REGION Network 83
   RUNG wire#powerrail
      Move(in := "Carrier_44_G120DControlWord", out1 => "DB402_SDC_CARRIER_DRIVE_DATA".Drive_Data.CARRIER[44].Drive_Control)
      Move(in := "Carrier_44_G120DStatusWord", out1 => "DB402_SDC_CARRIER_DRIVE_DATA".Drive_Data.CARRIER[44].Drive_Status)
   END_RUNG
   // the same network as SCL:
   "DB402_SDC_CARRIER_DRIVE_DATA".Drive_Data.CARRIER[44].Drive_Control := "Carrier_44_G120DControlWord";
   "DB402_SDC_CARRIER_DRIVE_DATA".Drive_Data.CARRIER[44].Drive_Status := "Carrier_44_G120DStatusWord";
END_REGION

REGION Network 84
   RUNG wire#powerrail
      Move(in := "Carrier_44_SDCFaultCode", out1 => "DB_SDC_EMS_TA".EMS[44].TA[1].FAULT)
      wire#w1
      Move(in := "Carrier_44_SDCFaultCode", out1 => "EMS".Carrier[44].SDC_IN.CarrierDriveFaults)
   END_RUNG
   RUNG wire#powerrail
      Contact( "IndiconTempDebugON" )
   END_RUNG wire#w1
   // the same network as SCL:
   "DB_SDC_EMS_TA".EMS[44].TA[1].FAULT := "Carrier_44_SDCFaultCode";
   IF TRUE OR "IndiconTempDebugON" THEN
       "EMS".Carrier[44].SDC_IN.CarrierDriveFaults := "Carrier_44_SDCFaultCode";
   END_IF;
END_REGION

REGION Network 85
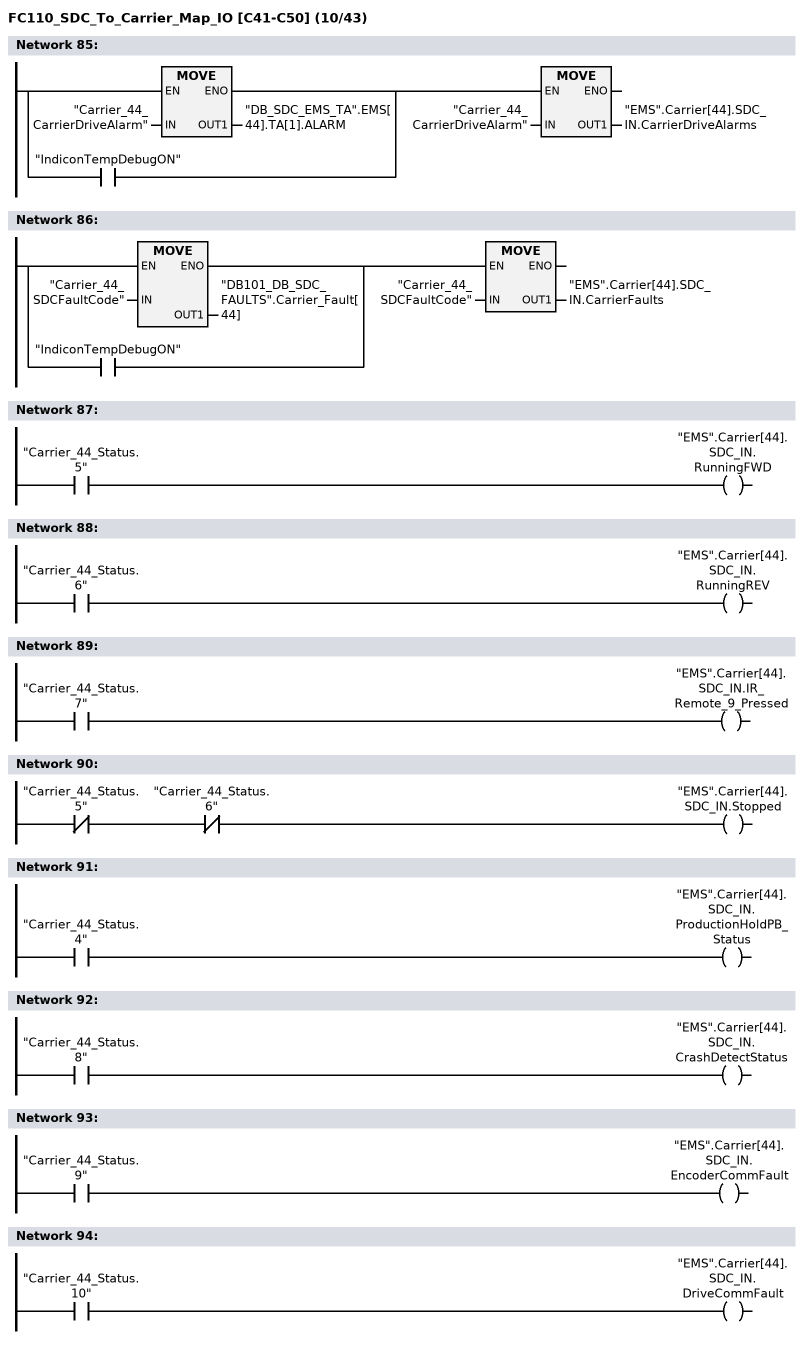
   RUNG wire#powerrail
      Move(in := "Carrier_44_CarrierDriveAlarm", out1 => "DB_SDC_EMS_TA".EMS[44].TA[1].ALARM)
      wire#w1
      Move(in := "Carrier_44_CarrierDriveAlarm", out1 => "EMS".Carrier[44].SDC_IN.CarrierDriveAlarms)
   END_RUNG
   RUNG wire#powerrail
      Contact( "IndiconTempDebugON" )
   END_RUNG wire#w1
   // the same network as SCL:
   "DB_SDC_EMS_TA".EMS[44].TA[1].ALARM := "Carrier_44_CarrierDriveAlarm";
   IF TRUE OR "IndiconTempDebugON" THEN
       "EMS".Carrier[44].SDC_IN.CarrierDriveAlarms := "Carrier_44_CarrierDriveAlarm";
   END_IF;
END_REGION

REGION Network 86
   RUNG wire#powerrail
      Move(in := "Carrier_44_SDCFaultCode", out1 => "DB101_DB_SDC_FAULTS".Carrier_Fault[44])
      wire#w1
      Move(in := "Carrier_44_SDCFaultCode", out1 => "EMS".Carrier[44].SDC_IN.CarrierFaults)
   END_RUNG
   RUNG wire#powerrail
      Contact( "IndiconTempDebugON" )
   END_RUNG wire#w1
   // the same network as SCL:
   "DB101_DB_SDC_FAULTS".Carrier_Fault[44] := "Carrier_44_SDCFaultCode";
   IF TRUE OR "IndiconTempDebugON" THEN
       "EMS".Carrier[44].SDC_IN.CarrierFaults := "Carrier_44_SDCFaultCode";
   END_IF;
END_REGION

REGION Network 87
   RUNG wire#powerrail
      Contact( "Carrier_44_Status.5" )
      Coil( "EMS".Carrier[44].SDC_IN.RunningFWD )
   END_RUNG
   // the same network as SCL:
   "EMS".Carrier[44].SDC_IN.RunningFWD := "Carrier_44_Status.5";
END_REGION

REGION Network 88
   RUNG wire#powerrail
      Contact( "Carrier_44_Status.6" )
      Coil( "EMS".Carrier[44].SDC_IN.RunningREV )
   END_RUNG
   // the same network as SCL:
   "EMS".Carrier[44].SDC_IN.RunningREV := "Carrier_44_Status.6";
END_REGION

REGION Network 89
   RUNG wire#powerrail
      Contact( "Carrier_44_Status.7" )
      Coil( "EMS".Carrier[44].SDC_IN.IR_Remote_9_Pressed )
   END_RUNG
   // the same network as SCL:
   "EMS".Carrier[44].SDC_IN.IR_Remote_9_Pressed := "Carrier_44_Status.7";
END_REGION

REGION Network 90
   RUNG wire#powerrail
      I_Contact( "Carrier_44_Status.5" )
      I_Contact( "Carrier_44_Status.6" )
      Coil( "EMS".Carrier[44].SDC_IN.Stopped )
   END_RUNG
   // the same network as SCL:
   "EMS".Carrier[44].SDC_IN.Stopped := NOT "Carrier_44_Status.5" AND NOT "Carrier_44_Status.6";
END_REGION

REGION Network 91
   RUNG wire#powerrail
      Contact( "Carrier_44_Status.4" )
      Coil( "EMS".Carrier[44].SDC_IN.ProductionHoldPB_Status )
   END_RUNG
   // the same network as SCL:
   "EMS".Carrier[44].SDC_IN.ProductionHoldPB_Status := "Carrier_44_Status.4";
END_REGION

REGION Network 92
   RUNG wire#powerrail
      Contact( "Carrier_44_Status.8" )
      Coil( "EMS".Carrier[44].SDC_IN.CrashDetectStatus )
   END_RUNG
   // the same network as SCL:
   "EMS".Carrier[44].SDC_IN.CrashDetectStatus := "Carrier_44_Status.8";
END_REGION

REGION Network 93
   RUNG wire#powerrail
      Contact( "Carrier_44_Status.9" )
      Coil( "EMS".Carrier[44].SDC_IN.EncoderCommFault )
   END_RUNG
   // the same network as SCL:
   "EMS".Carrier[44].SDC_IN.EncoderCommFault := "Carrier_44_Status.9";
END_REGION

REGION Network 94
   RUNG wire#powerrail
      Contact( "Carrier_44_Status.10" )
      Coil( "EMS".Carrier[44].SDC_IN.DriveCommFault )
   END_RUNG
   // the same network as SCL:
   "EMS".Carrier[44].SDC_IN.DriveCommFault := "Carrier_44_Status.10";
END_REGION

REGION Network 95
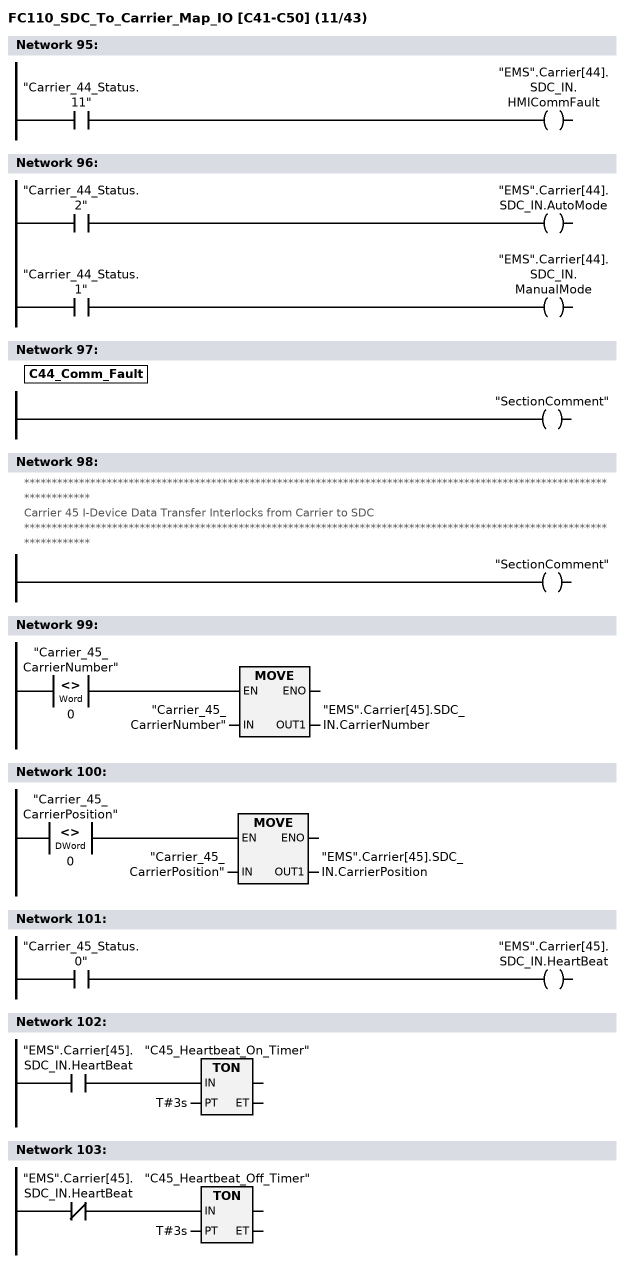
   RUNG wire#powerrail
      Contact( "Carrier_44_Status.11" )
      Coil( "EMS".Carrier[44].SDC_IN.HMICommFault )
   END_RUNG
   // the same network as SCL:
   "EMS".Carrier[44].SDC_IN.HMICommFault := "Carrier_44_Status.11";
END_REGION

REGION Network 96
   RUNG wire#powerrail
      Contact( "Carrier_44_Status.2" )
      Coil( "EMS".Carrier[44].SDC_IN.AutoMode )
   END_RUNG
   RUNG wire#powerrail
      Contact( "Carrier_44_Status.1" )
      Coil( "EMS".Carrier[44].SDC_IN.ManualMode )
   END_RUNG
   // the same network as SCL:
   "EMS".Carrier[44].SDC_IN.AutoMode := "Carrier_44_Status.2";
   "EMS".Carrier[44].SDC_IN.ManualMode := "Carrier_44_Status.1";
END_REGION

REGION Network 97
   Label( C44_Comm_Fault )
   RUNG wire#powerrail
      Coil( "SectionComment" )
   END_RUNG
   // the same network as SCL:
   C44_Comm_Fault:
   "SectionComment" := TRUE;
END_REGION

REGION Network 98
   // **********************************************************************************************************************
   // 
   // Carrier 45 I-Device Data Transfer Interlocks from Carrier to SDC
   // 
   // **********************************************************************************************************************
   RUNG wire#powerrail
      Coil( "SectionComment" )
   END_RUNG
   // the same network as SCL:
   "SectionComment" := TRUE;
END_REGION

REGION Network 99
   RUNG wire#powerrail
      { S7_Templates := "SrcType := Word" } NE_Contact(in1 := "Carrier_45_CarrierNumber", in2 := 0)
      Move(in := "Carrier_45_CarrierNumber", out1 => "EMS".Carrier[45].SDC_IN.CarrierNumber)
   END_RUNG
   // the same network as SCL:
   IF "Carrier_45_CarrierNumber" <> 0 THEN
       "EMS".Carrier[45].SDC_IN.CarrierNumber := "Carrier_45_CarrierNumber";
   END_IF;
END_REGION

REGION Network 100
   RUNG wire#powerrail
      { S7_Templates := "SrcType := DWord" } NE_Contact(in1 := "Carrier_45_CarrierPosition", in2 := 0)
      Move(in := "Carrier_45_CarrierPosition", out1 => "EMS".Carrier[45].SDC_IN.CarrierPosition)
   END_RUNG
   // the same network as SCL:
   IF "Carrier_45_CarrierPosition" <> 0 THEN
       "EMS".Carrier[45].SDC_IN.CarrierPosition := "Carrier_45_CarrierPosition";
   END_IF;
END_REGION

REGION Network 101
   RUNG wire#powerrail
      Contact( "Carrier_45_Status.0" )
      Coil( "EMS".Carrier[45].SDC_IN.HeartBeat )
   END_RUNG
   // the same network as SCL:
   "EMS".Carrier[45].SDC_IN.HeartBeat := "Carrier_45_Status.0";
END_REGION

REGION Network 102
   "C45_Heartbeat_On_Timer".TON(IN := "EMS".Carrier[45].SDC_IN.HeartBeat, PT := T#3s);
END_REGION

REGION Network 103
   "C45_Heartbeat_Off_Timer".TON(IN := NOT "EMS".Carrier[45].SDC_IN.HeartBeat, PT := T#3s);
END_REGION

REGION Network 104
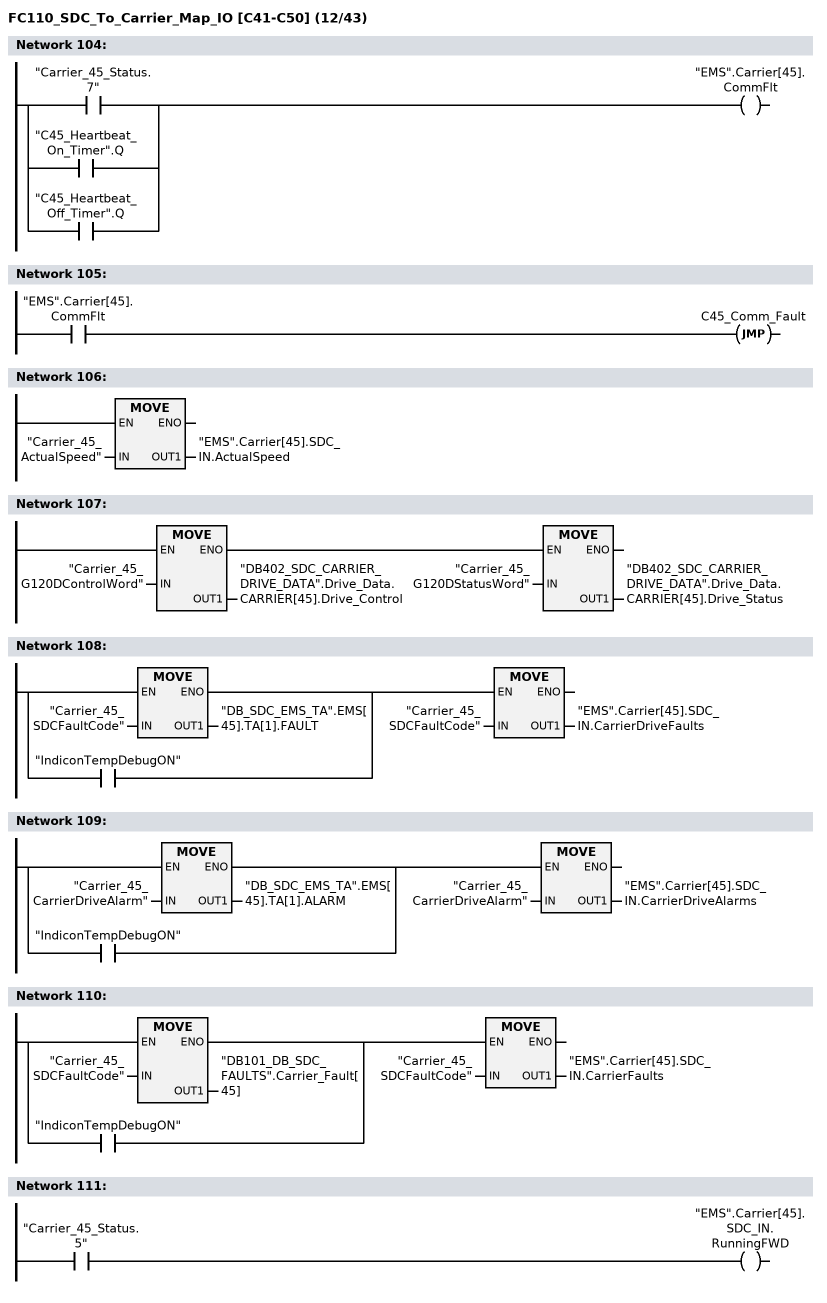
   RUNG wire#powerrail
      Contact( "Carrier_45_Status.7" )
      wire#w1
      Coil( "EMS".Carrier[45].CommFlt )
   END_RUNG
   RUNG wire#powerrail
      Contact( "C45_Heartbeat_On_Timer".Q )
   END_RUNG wire#w1
   RUNG wire#powerrail
      Contact( "C45_Heartbeat_Off_Timer".Q )
   END_RUNG wire#w1
   // the same network as SCL:
   "EMS".Carrier[45].CommFlt := "Carrier_45_Status.7" OR "C45_Heartbeat_On_Timer".Q OR "C45_Heartbeat_Off_Timer".Q;
END_REGION

REGION Network 105
   RUNG wire#powerrail
      Contact( "EMS".Carrier[45].CommFlt )
      JumpCoil( C45_Comm_Fault )
   END_RUNG
   // the same network as SCL:
   IF "EMS".Carrier[45].CommFlt THEN GOTO C45_Comm_Fault; END_IF;
END_REGION

REGION Network 106
   RUNG wire#powerrail
      Move(in := "Carrier_45_ActualSpeed", out1 => "EMS".Carrier[45].SDC_IN.ActualSpeed)
   END_RUNG
   // the same network as SCL:
   "EMS".Carrier[45].SDC_IN.ActualSpeed := "Carrier_45_ActualSpeed";
END_REGION

REGION Network 107
   RUNG wire#powerrail
      Move(in := "Carrier_45_G120DControlWord", out1 => "DB402_SDC_CARRIER_DRIVE_DATA".Drive_Data.CARRIER[45].Drive_Control)
      Move(in := "Carrier_45_G120DStatusWord", out1 => "DB402_SDC_CARRIER_DRIVE_DATA".Drive_Data.CARRIER[45].Drive_Status)
   END_RUNG
   // the same network as SCL:
   "DB402_SDC_CARRIER_DRIVE_DATA".Drive_Data.CARRIER[45].Drive_Control := "Carrier_45_G120DControlWord";
   "DB402_SDC_CARRIER_DRIVE_DATA".Drive_Data.CARRIER[45].Drive_Status := "Carrier_45_G120DStatusWord";
END_REGION

REGION Network 108
   RUNG wire#powerrail
      Move(in := "Carrier_45_SDCFaultCode", out1 => "DB_SDC_EMS_TA".EMS[45].TA[1].FAULT)
      wire#w1
      Move(in := "Carrier_45_SDCFaultCode", out1 => "EMS".Carrier[45].SDC_IN.CarrierDriveFaults)
   END_RUNG
   RUNG wire#powerrail
      Contact( "IndiconTempDebugON" )
   END_RUNG wire#w1
   // the same network as SCL:
   "DB_SDC_EMS_TA".EMS[45].TA[1].FAULT := "Carrier_45_SDCFaultCode";
   IF TRUE OR "IndiconTempDebugON" THEN
       "EMS".Carrier[45].SDC_IN.CarrierDriveFaults := "Carrier_45_SDCFaultCode";
   END_IF;
END_REGION

REGION Network 109
   RUNG wire#powerrail
      Move(in := "Carrier_45_CarrierDriveAlarm", out1 => "DB_SDC_EMS_TA".EMS[45].TA[1].ALARM)
      wire#w1
      Move(in := "Carrier_45_CarrierDriveAlarm", out1 => "EMS".Carrier[45].SDC_IN.CarrierDriveAlarms)
   END_RUNG
   RUNG wire#powerrail
      Contact( "IndiconTempDebugON" )
   END_RUNG wire#w1
   // the same network as SCL:
   "DB_SDC_EMS_TA".EMS[45].TA[1].ALARM := "Carrier_45_CarrierDriveAlarm";
   IF TRUE OR "IndiconTempDebugON" THEN
       "EMS".Carrier[45].SDC_IN.CarrierDriveAlarms := "Carrier_45_CarrierDriveAlarm";
   END_IF;
END_REGION

REGION Network 110
   RUNG wire#powerrail
      Move(in := "Carrier_45_SDCFaultCode", out1 => "DB101_DB_SDC_FAULTS".Carrier_Fault[45])
      wire#w1
      Move(in := "Carrier_45_SDCFaultCode", out1 => "EMS".Carrier[45].SDC_IN.CarrierFaults)
   END_RUNG
   RUNG wire#powerrail
      Contact( "IndiconTempDebugON" )
   END_RUNG wire#w1
   // the same network as SCL:
   "DB101_DB_SDC_FAULTS".Carrier_Fault[45] := "Carrier_45_SDCFaultCode";
   IF TRUE OR "IndiconTempDebugON" THEN
       "EMS".Carrier[45].SDC_IN.CarrierFaults := "Carrier_45_SDCFaultCode";
   END_IF;
END_REGION

REGION Network 111
   RUNG wire#powerrail
      Contact( "Carrier_45_Status.5" )
      Coil( "EMS".Carrier[45].SDC_IN.RunningFWD )
   END_RUNG
   // the same network as SCL:
   "EMS".Carrier[45].SDC_IN.RunningFWD := "Carrier_45_Status.5";
END_REGION

REGION Network 112
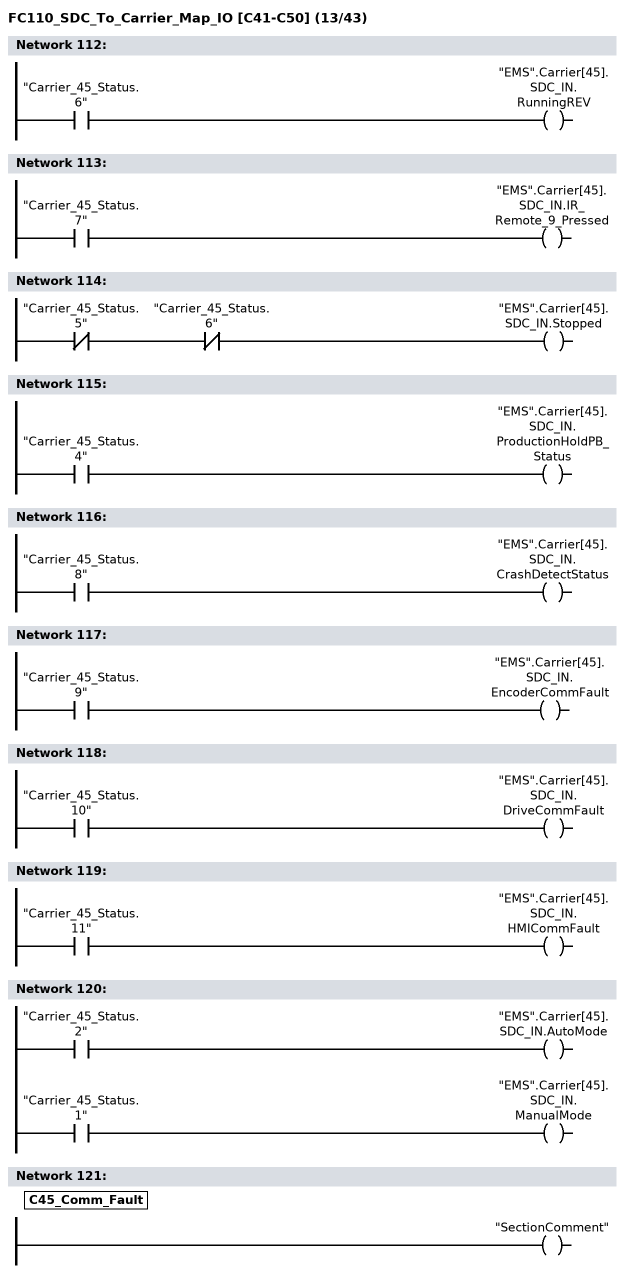
   RUNG wire#powerrail
      Contact( "Carrier_45_Status.6" )
      Coil( "EMS".Carrier[45].SDC_IN.RunningREV )
   END_RUNG
   // the same network as SCL:
   "EMS".Carrier[45].SDC_IN.RunningREV := "Carrier_45_Status.6";
END_REGION

REGION Network 113
   RUNG wire#powerrail
      Contact( "Carrier_45_Status.7" )
      Coil( "EMS".Carrier[45].SDC_IN.IR_Remote_9_Pressed )
   END_RUNG
   // the same network as SCL:
   "EMS".Carrier[45].SDC_IN.IR_Remote_9_Pressed := "Carrier_45_Status.7";
END_REGION

REGION Network 114
   RUNG wire#powerrail
      I_Contact( "Carrier_45_Status.5" )
      I_Contact( "Carrier_45_Status.6" )
      Coil( "EMS".Carrier[45].SDC_IN.Stopped )
   END_RUNG
   // the same network as SCL:
   "EMS".Carrier[45].SDC_IN.Stopped := NOT "Carrier_45_Status.5" AND NOT "Carrier_45_Status.6";
END_REGION

REGION Network 115
   RUNG wire#powerrail
      Contact( "Carrier_45_Status.4" )
      Coil( "EMS".Carrier[45].SDC_IN.ProductionHoldPB_Status )
   END_RUNG
   // the same network as SCL:
   "EMS".Carrier[45].SDC_IN.ProductionHoldPB_Status := "Carrier_45_Status.4";
END_REGION

REGION Network 116
   RUNG wire#powerrail
      Contact( "Carrier_45_Status.8" )
      Coil( "EMS".Carrier[45].SDC_IN.CrashDetectStatus )
   END_RUNG
   // the same network as SCL:
   "EMS".Carrier[45].SDC_IN.CrashDetectStatus := "Carrier_45_Status.8";
END_REGION

REGION Network 117
   RUNG wire#powerrail
      Contact( "Carrier_45_Status.9" )
      Coil( "EMS".Carrier[45].SDC_IN.EncoderCommFault )
   END_RUNG
   // the same network as SCL:
   "EMS".Carrier[45].SDC_IN.EncoderCommFault := "Carrier_45_Status.9";
END_REGION

REGION Network 118
   RUNG wire#powerrail
      Contact( "Carrier_45_Status.10" )
      Coil( "EMS".Carrier[45].SDC_IN.DriveCommFault )
   END_RUNG
   // the same network as SCL:
   "EMS".Carrier[45].SDC_IN.DriveCommFault := "Carrier_45_Status.10";
END_REGION

REGION Network 119
   RUNG wire#powerrail
      Contact( "Carrier_45_Status.11" )
      Coil( "EMS".Carrier[45].SDC_IN.HMICommFault )
   END_RUNG
   // the same network as SCL:
   "EMS".Carrier[45].SDC_IN.HMICommFault := "Carrier_45_Status.11";
END_REGION

REGION Network 120
   RUNG wire#powerrail
      Contact( "Carrier_45_Status.2" )
      Coil( "EMS".Carrier[45].SDC_IN.AutoMode )
   END_RUNG
   RUNG wire#powerrail
      Contact( "Carrier_45_Status.1" )
      Coil( "EMS".Carrier[45].SDC_IN.ManualMode )
   END_RUNG
   // the same network as SCL:
   "EMS".Carrier[45].SDC_IN.AutoMode := "Carrier_45_Status.2";
   "EMS".Carrier[45].SDC_IN.ManualMode := "Carrier_45_Status.1";
END_REGION

REGION Network 121
   Label( C45_Comm_Fault )
   RUNG wire#powerrail
      Coil( "SectionComment" )
   END_RUNG
   // the same network as SCL:
   C45_Comm_Fault:
   "SectionComment" := TRUE;
END_REGION

REGION Network 122
   // **********************************************************************************************************************
   // 
   // Carrier 46 I-Device Data Transfer Interlocks from Carrier to SDC
   // 
   // **********************************************************************************************************************
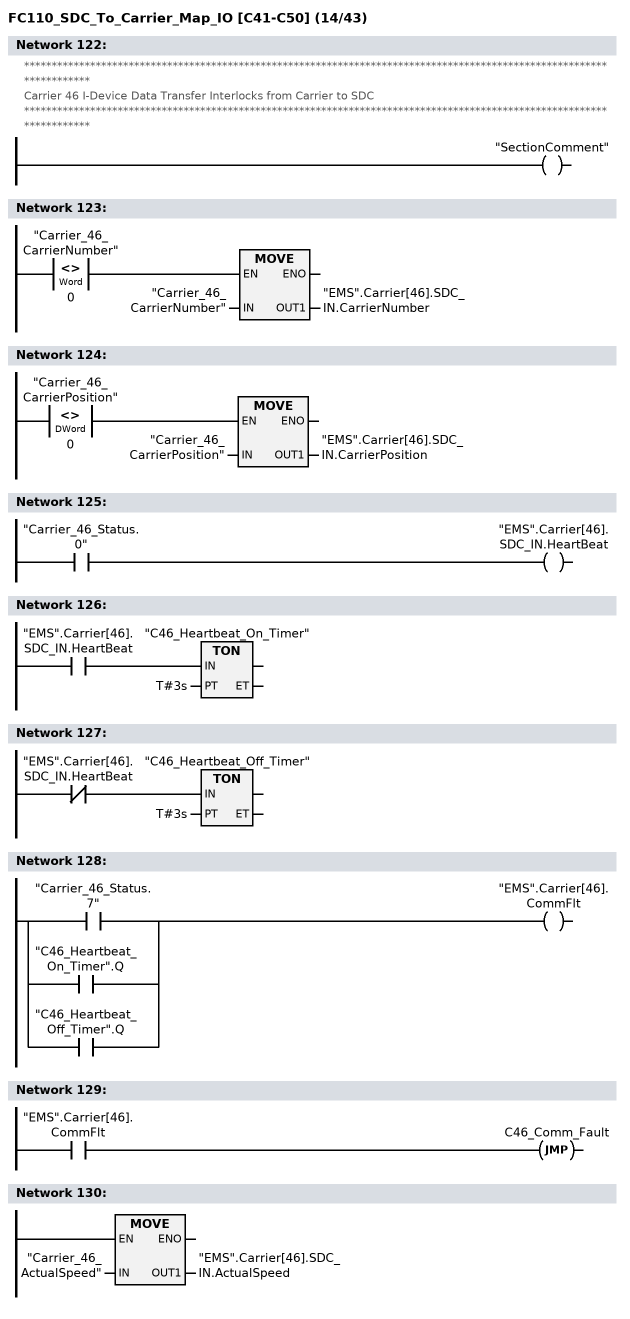
   RUNG wire#powerrail
      Coil( "SectionComment" )
   END_RUNG
   // the same network as SCL:
   "SectionComment" := TRUE;
END_REGION

REGION Network 123
   RUNG wire#powerrail
      { S7_Templates := "SrcType := Word" } NE_Contact(in1 := "Carrier_46_CarrierNumber", in2 := 0)
      Move(in := "Carrier_46_CarrierNumber", out1 => "EMS".Carrier[46].SDC_IN.CarrierNumber)
   END_RUNG
   // the same network as SCL:
   IF "Carrier_46_CarrierNumber" <> 0 THEN
       "EMS".Carrier[46].SDC_IN.CarrierNumber := "Carrier_46_CarrierNumber";
   END_IF;
END_REGION

REGION Network 124
   RUNG wire#powerrail
      { S7_Templates := "SrcType := DWord" } NE_Contact(in1 := "Carrier_46_CarrierPosition", in2 := 0)
      Move(in := "Carrier_46_CarrierPosition", out1 => "EMS".Carrier[46].SDC_IN.CarrierPosition)
   END_RUNG
   // the same network as SCL:
   IF "Carrier_46_CarrierPosition" <> 0 THEN
       "EMS".Carrier[46].SDC_IN.CarrierPosition := "Carrier_46_CarrierPosition";
   END_IF;
END_REGION

REGION Network 125
   RUNG wire#powerrail
      Contact( "Carrier_46_Status.0" )
      Coil( "EMS".Carrier[46].SDC_IN.HeartBeat )
   END_RUNG
   // the same network as SCL:
   "EMS".Carrier[46].SDC_IN.HeartBeat := "Carrier_46_Status.0";
END_REGION

REGION Network 126
   "C46_Heartbeat_On_Timer".TON(IN := "EMS".Carrier[46].SDC_IN.HeartBeat, PT := T#3s);
END_REGION

REGION Network 127
   "C46_Heartbeat_Off_Timer".TON(IN := NOT "EMS".Carrier[46].SDC_IN.HeartBeat, PT := T#3s);
END_REGION

REGION Network 128
   RUNG wire#powerrail
      Contact( "Carrier_46_Status.7" )
      wire#w1
      Coil( "EMS".Carrier[46].CommFlt )
   END_RUNG
   RUNG wire#powerrail
      Contact( "C46_Heartbeat_On_Timer".Q )
   END_RUNG wire#w1
   RUNG wire#powerrail
      Contact( "C46_Heartbeat_Off_Timer".Q )
   END_RUNG wire#w1
   // the same network as SCL:
   "EMS".Carrier[46].CommFlt := "Carrier_46_Status.7" OR "C46_Heartbeat_On_Timer".Q OR "C46_Heartbeat_Off_Timer".Q;
END_REGION

REGION Network 129
   RUNG wire#powerrail
      Contact( "EMS".Carrier[46].CommFlt )
      JumpCoil( C46_Comm_Fault )
   END_RUNG
   // the same network as SCL:
   IF "EMS".Carrier[46].CommFlt THEN GOTO C46_Comm_Fault; END_IF;
END_REGION

REGION Network 130
   RUNG wire#powerrail
      Move(in := "Carrier_46_ActualSpeed", out1 => "EMS".Carrier[46].SDC_IN.ActualSpeed)
   END_RUNG
   // the same network as SCL:
   "EMS".Carrier[46].SDC_IN.ActualSpeed := "Carrier_46_ActualSpeed";
END_REGION

REGION Network 131
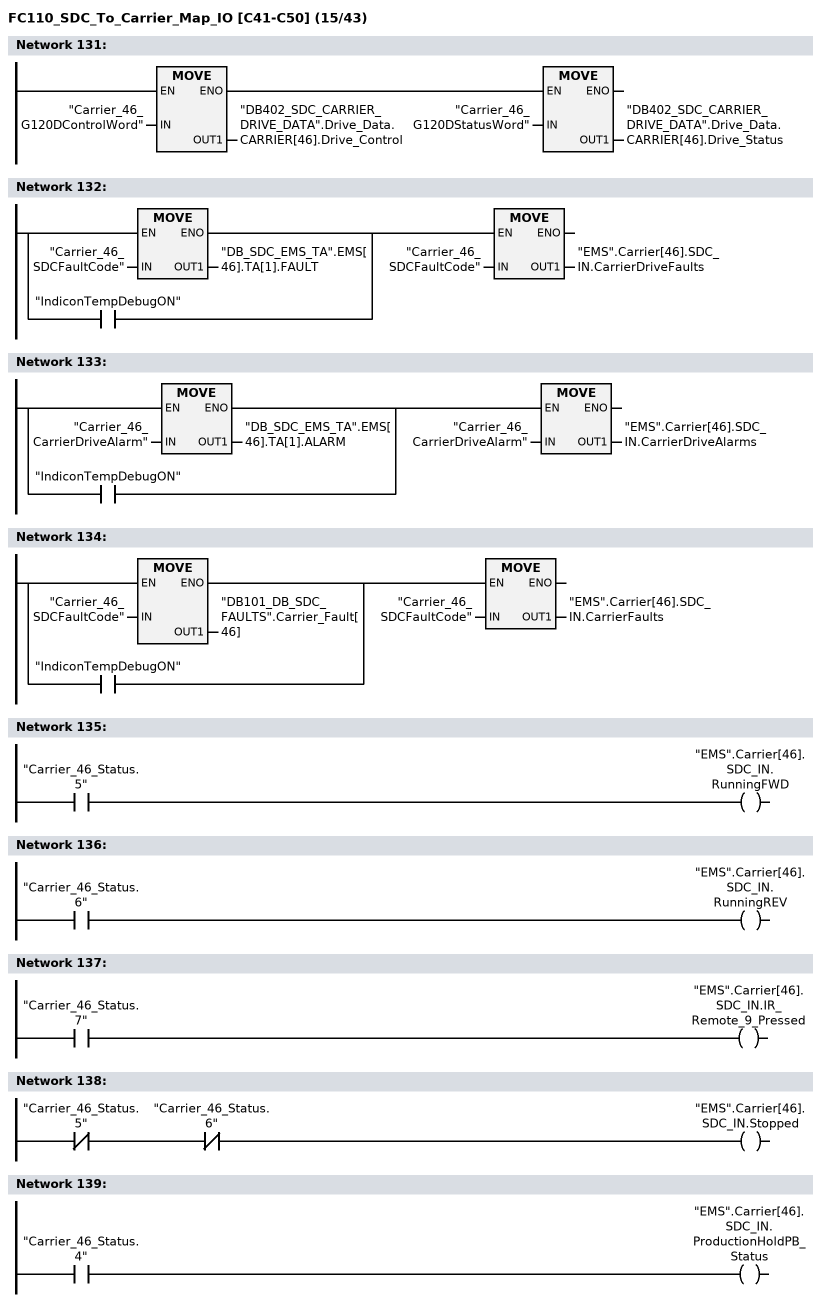
   RUNG wire#powerrail
      Move(in := "Carrier_46_G120DControlWord", out1 => "DB402_SDC_CARRIER_DRIVE_DATA".Drive_Data.CARRIER[46].Drive_Control)
      Move(in := "Carrier_46_G120DStatusWord", out1 => "DB402_SDC_CARRIER_DRIVE_DATA".Drive_Data.CARRIER[46].Drive_Status)
   END_RUNG
   // the same network as SCL:
   "DB402_SDC_CARRIER_DRIVE_DATA".Drive_Data.CARRIER[46].Drive_Control := "Carrier_46_G120DControlWord";
   "DB402_SDC_CARRIER_DRIVE_DATA".Drive_Data.CARRIER[46].Drive_Status := "Carrier_46_G120DStatusWord";
END_REGION

REGION Network 132
   RUNG wire#powerrail
      Move(in := "Carrier_46_SDCFaultCode", out1 => "DB_SDC_EMS_TA".EMS[46].TA[1].FAULT)
      wire#w1
      Move(in := "Carrier_46_SDCFaultCode", out1 => "EMS".Carrier[46].SDC_IN.CarrierDriveFaults)
   END_RUNG
   RUNG wire#powerrail
      Contact( "IndiconTempDebugON" )
   END_RUNG wire#w1
   // the same network as SCL:
   "DB_SDC_EMS_TA".EMS[46].TA[1].FAULT := "Carrier_46_SDCFaultCode";
   IF TRUE OR "IndiconTempDebugON" THEN
       "EMS".Carrier[46].SDC_IN.CarrierDriveFaults := "Carrier_46_SDCFaultCode";
   END_IF;
END_REGION

REGION Network 133
   RUNG wire#powerrail
      Move(in := "Carrier_46_CarrierDriveAlarm", out1 => "DB_SDC_EMS_TA".EMS[46].TA[1].ALARM)
      wire#w1
      Move(in := "Carrier_46_CarrierDriveAlarm", out1 => "EMS".Carrier[46].SDC_IN.CarrierDriveAlarms)
   END_RUNG
   RUNG wire#powerrail
      Contact( "IndiconTempDebugON" )
   END_RUNG wire#w1
   // the same network as SCL:
   "DB_SDC_EMS_TA".EMS[46].TA[1].ALARM := "Carrier_46_CarrierDriveAlarm";
   IF TRUE OR "IndiconTempDebugON" THEN
       "EMS".Carrier[46].SDC_IN.CarrierDriveAlarms := "Carrier_46_CarrierDriveAlarm";
   END_IF;
END_REGION

REGION Network 134
   RUNG wire#powerrail
      Move(in := "Carrier_46_SDCFaultCode", out1 => "DB101_DB_SDC_FAULTS".Carrier_Fault[46])
      wire#w1
      Move(in := "Carrier_46_SDCFaultCode", out1 => "EMS".Carrier[46].SDC_IN.CarrierFaults)
   END_RUNG
   RUNG wire#powerrail
      Contact( "IndiconTempDebugON" )
   END_RUNG wire#w1
   // the same network as SCL:
   "DB101_DB_SDC_FAULTS".Carrier_Fault[46] := "Carrier_46_SDCFaultCode";
   IF TRUE OR "IndiconTempDebugON" THEN
       "EMS".Carrier[46].SDC_IN.CarrierFaults := "Carrier_46_SDCFaultCode";
   END_IF;
END_REGION

REGION Network 135
   RUNG wire#powerrail
      Contact( "Carrier_46_Status.5" )
      Coil( "EMS".Carrier[46].SDC_IN.RunningFWD )
   END_RUNG
   // the same network as SCL:
   "EMS".Carrier[46].SDC_IN.RunningFWD := "Carrier_46_Status.5";
END_REGION

REGION Network 136
   RUNG wire#powerrail
      Contact( "Carrier_46_Status.6" )
      Coil( "EMS".Carrier[46].SDC_IN.RunningREV )
   END_RUNG
   // the same network as SCL:
   "EMS".Carrier[46].SDC_IN.RunningREV := "Carrier_46_Status.6";
END_REGION

REGION Network 137
   RUNG wire#powerrail
      Contact( "Carrier_46_Status.7" )
      Coil( "EMS".Carrier[46].SDC_IN.IR_Remote_9_Pressed )
   END_RUNG
   // the same network as SCL:
   "EMS".Carrier[46].SDC_IN.IR_Remote_9_Pressed := "Carrier_46_Status.7";
END_REGION

REGION Network 138
   RUNG wire#powerrail
      I_Contact( "Carrier_46_Status.5" )
      I_Contact( "Carrier_46_Status.6" )
      Coil( "EMS".Carrier[46].SDC_IN.Stopped )
   END_RUNG
   // the same network as SCL:
   "EMS".Carrier[46].SDC_IN.Stopped := NOT "Carrier_46_Status.5" AND NOT "Carrier_46_Status.6";
END_REGION

REGION Network 139
   RUNG wire#powerrail
      Contact( "Carrier_46_Status.4" )
      Coil( "EMS".Carrier[46].SDC_IN.ProductionHoldPB_Status )
   END_RUNG
   // the same network as SCL:
   "EMS".Carrier[46].SDC_IN.ProductionHoldPB_Status := "Carrier_46_Status.4";
END_REGION

REGION Network 140
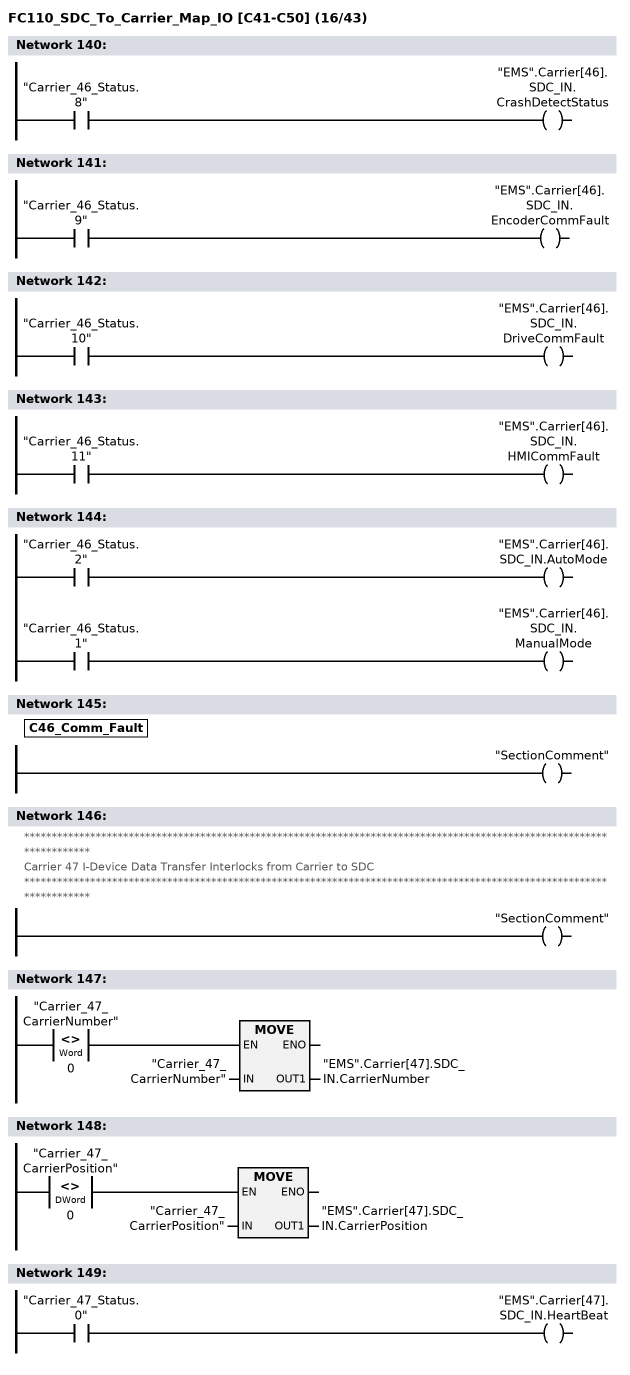
   RUNG wire#powerrail
      Contact( "Carrier_46_Status.8" )
      Coil( "EMS".Carrier[46].SDC_IN.CrashDetectStatus )
   END_RUNG
   // the same network as SCL:
   "EMS".Carrier[46].SDC_IN.CrashDetectStatus := "Carrier_46_Status.8";
END_REGION

REGION Network 141
   RUNG wire#powerrail
      Contact( "Carrier_46_Status.9" )
      Coil( "EMS".Carrier[46].SDC_IN.EncoderCommFault )
   END_RUNG
   // the same network as SCL:
   "EMS".Carrier[46].SDC_IN.EncoderCommFault := "Carrier_46_Status.9";
END_REGION

REGION Network 142
   RUNG wire#powerrail
      Contact( "Carrier_46_Status.10" )
      Coil( "EMS".Carrier[46].SDC_IN.DriveCommFault )
   END_RUNG
   // the same network as SCL:
   "EMS".Carrier[46].SDC_IN.DriveCommFault := "Carrier_46_Status.10";
END_REGION

REGION Network 143
   RUNG wire#powerrail
      Contact( "Carrier_46_Status.11" )
      Coil( "EMS".Carrier[46].SDC_IN.HMICommFault )
   END_RUNG
   // the same network as SCL:
   "EMS".Carrier[46].SDC_IN.HMICommFault := "Carrier_46_Status.11";
END_REGION

REGION Network 144
   RUNG wire#powerrail
      Contact( "Carrier_46_Status.2" )
      Coil( "EMS".Carrier[46].SDC_IN.AutoMode )
   END_RUNG
   RUNG wire#powerrail
      Contact( "Carrier_46_Status.1" )
      Coil( "EMS".Carrier[46].SDC_IN.ManualMode )
   END_RUNG
   // the same network as SCL:
   "EMS".Carrier[46].SDC_IN.AutoMode := "Carrier_46_Status.2";
   "EMS".Carrier[46].SDC_IN.ManualMode := "Carrier_46_Status.1";
END_REGION

REGION Network 145
   Label( C46_Comm_Fault )
   RUNG wire#powerrail
      Coil( "SectionComment" )
   END_RUNG
   // the same network as SCL:
   C46_Comm_Fault:
   "SectionComment" := TRUE;
END_REGION

REGION Network 146
   // **********************************************************************************************************************
   // 
   // Carrier 47 I-Device Data Transfer Interlocks from Carrier to SDC
   // 
   // **********************************************************************************************************************
   RUNG wire#powerrail
      Coil( "SectionComment" )
   END_RUNG
   // the same network as SCL:
   "SectionComment" := TRUE;
END_REGION

REGION Network 147
   RUNG wire#powerrail
      { S7_Templates := "SrcType := Word" } NE_Contact(in1 := "Carrier_47_CarrierNumber", in2 := 0)
      Move(in := "Carrier_47_CarrierNumber", out1 => "EMS".Carrier[47].SDC_IN.CarrierNumber)
   END_RUNG
   // the same network as SCL:
   IF "Carrier_47_CarrierNumber" <> 0 THEN
       "EMS".Carrier[47].SDC_IN.CarrierNumber := "Carrier_47_CarrierNumber";
   END_IF;
END_REGION

REGION Network 148
   RUNG wire#powerrail
      { S7_Templates := "SrcType := DWord" } NE_Contact(in1 := "Carrier_47_CarrierPosition", in2 := 0)
      Move(in := "Carrier_47_CarrierPosition", out1 => "EMS".Carrier[47].SDC_IN.CarrierPosition)
   END_RUNG
   // the same network as SCL:
   IF "Carrier_47_CarrierPosition" <> 0 THEN
       "EMS".Carrier[47].SDC_IN.CarrierPosition := "Carrier_47_CarrierPosition";
   END_IF;
END_REGION

REGION Network 149
   RUNG wire#powerrail
      Contact( "Carrier_47_Status.0" )
      Coil( "EMS".Carrier[47].SDC_IN.HeartBeat )
   END_RUNG
   // the same network as SCL:
   "EMS".Carrier[47].SDC_IN.HeartBeat := "Carrier_47_Status.0";
END_REGION

REGION Network 150
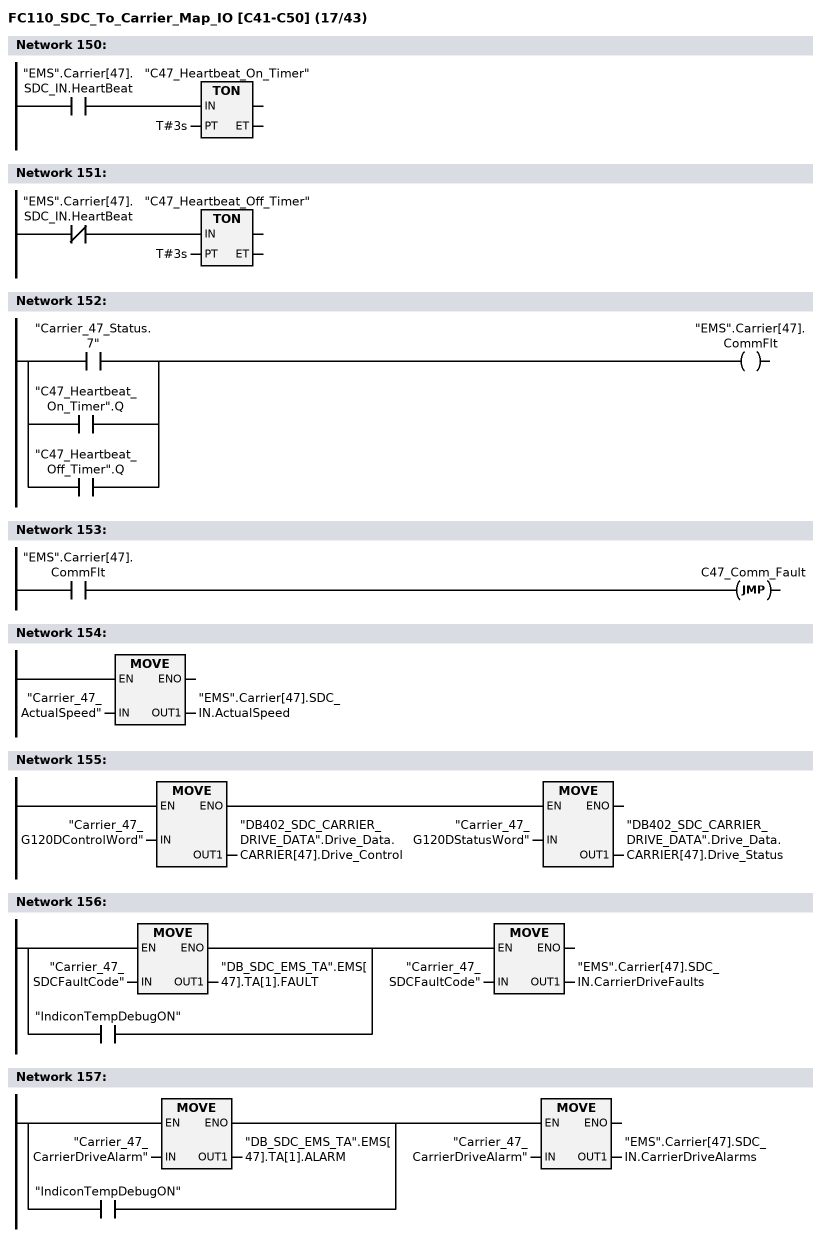
   "C47_Heartbeat_On_Timer".TON(IN := "EMS".Carrier[47].SDC_IN.HeartBeat, PT := T#3s);
END_REGION

REGION Network 151
   "C47_Heartbeat_Off_Timer".TON(IN := NOT "EMS".Carrier[47].SDC_IN.HeartBeat, PT := T#3s);
END_REGION

REGION Network 152
   RUNG wire#powerrail
      Contact( "Carrier_47_Status.7" )
      wire#w1
      Coil( "EMS".Carrier[47].CommFlt )
   END_RUNG
   RUNG wire#powerrail
      Contact( "C47_Heartbeat_On_Timer".Q )
   END_RUNG wire#w1
   RUNG wire#powerrail
      Contact( "C47_Heartbeat_Off_Timer".Q )
   END_RUNG wire#w1
   // the same network as SCL:
   "EMS".Carrier[47].CommFlt := "Carrier_47_Status.7" OR "C47_Heartbeat_On_Timer".Q OR "C47_Heartbeat_Off_Timer".Q;
END_REGION

REGION Network 153
   RUNG wire#powerrail
      Contact( "EMS".Carrier[47].CommFlt )
      JumpCoil( C47_Comm_Fault )
   END_RUNG
   // the same network as SCL:
   IF "EMS".Carrier[47].CommFlt THEN GOTO C47_Comm_Fault; END_IF;
END_REGION

REGION Network 154
   RUNG wire#powerrail
      Move(in := "Carrier_47_ActualSpeed", out1 => "EMS".Carrier[47].SDC_IN.ActualSpeed)
   END_RUNG
   // the same network as SCL:
   "EMS".Carrier[47].SDC_IN.ActualSpeed := "Carrier_47_ActualSpeed";
END_REGION

REGION Network 155
   RUNG wire#powerrail
      Move(in := "Carrier_47_G120DControlWord", out1 => "DB402_SDC_CARRIER_DRIVE_DATA".Drive_Data.CARRIER[47].Drive_Control)
      Move(in := "Carrier_47_G120DStatusWord", out1 => "DB402_SDC_CARRIER_DRIVE_DATA".Drive_Data.CARRIER[47].Drive_Status)
   END_RUNG
   // the same network as SCL:
   "DB402_SDC_CARRIER_DRIVE_DATA".Drive_Data.CARRIER[47].Drive_Control := "Carrier_47_G120DControlWord";
   "DB402_SDC_CARRIER_DRIVE_DATA".Drive_Data.CARRIER[47].Drive_Status := "Carrier_47_G120DStatusWord";
END_REGION

REGION Network 156
   RUNG wire#powerrail
      Move(in := "Carrier_47_SDCFaultCode", out1 => "DB_SDC_EMS_TA".EMS[47].TA[1].FAULT)
      wire#w1
      Move(in := "Carrier_47_SDCFaultCode", out1 => "EMS".Carrier[47].SDC_IN.CarrierDriveFaults)
   END_RUNG
   RUNG wire#powerrail
      Contact( "IndiconTempDebugON" )
   END_RUNG wire#w1
   // the same network as SCL:
   "DB_SDC_EMS_TA".EMS[47].TA[1].FAULT := "Carrier_47_SDCFaultCode";
   IF TRUE OR "IndiconTempDebugON" THEN
       "EMS".Carrier[47].SDC_IN.CarrierDriveFaults := "Carrier_47_SDCFaultCode";
   END_IF;
END_REGION

REGION Network 157
   RUNG wire#powerrail
      Move(in := "Carrier_47_CarrierDriveAlarm", out1 => "DB_SDC_EMS_TA".EMS[47].TA[1].ALARM)
      wire#w1
      Move(in := "Carrier_47_CarrierDriveAlarm", out1 => "EMS".Carrier[47].SDC_IN.CarrierDriveAlarms)
   END_RUNG
   RUNG wire#powerrail
      Contact( "IndiconTempDebugON" )
   END_RUNG wire#w1
   // the same network as SCL:
   "DB_SDC_EMS_TA".EMS[47].TA[1].ALARM := "Carrier_47_CarrierDriveAlarm";
   IF TRUE OR "IndiconTempDebugON" THEN
       "EMS".Carrier[47].SDC_IN.CarrierDriveAlarms := "Carrier_47_CarrierDriveAlarm";
   END_IF;
END_REGION

REGION Network 158
